REGION Network 5
   RUNG wire#powerrail
      { S7_Templates := "SrcType := Int" } EQ_Contact(in1 := #"BUFFER STATE", in2 := 0)
      I_Contact( #processing )
      I_Contact( #"MACHINE EXIT SENSOR" )
      I_Contact( #BUFFER_ITEMS_COUNT.QU )
      Move(in := 10, out1 => #"BUFFER STATE")
   END_RUNG
   // the same network as SCL:
   IF (#"BUFFER STATE" = 0) AND NOT #processing AND NOT #"MACHINE EXIT SENSOR" AND NOT #BUFFER_ITEMS_COUNT.QU THEN
       #"BUFFER STATE" := 10;
   END_IF;
END_REGION

REGION Network 6
   RUNG wire#powerrail
      #"ZONE 3 STOP BLADES LOGIC_Instance"("BUFFER STATE" := #"BUFFER STATE", "UP ELEVATOR STOP BLADE" => #"UP ELEVATOR STOP BLADE", "DOWN ELEVATOR STOP BLADE" => #"DOWN ELEVATOR STOP BLADE", "BRIDGE STOP BLADE 1" => #"BRIDGE STOP BLADE 1", "BRIDGE STOP BLADE 2" => #"BRIDGE STOP BLADE 2")
   END_RUNG
   // the same network as SCL:
   #"ZONE 3 STOP BLADES LOGIC_Instance"("BUFFER STATE" := #"BUFFER STATE",   // "ZONE 3 STOP BLADES LOGIC"
                           "UP ELEVATOR STOP BLADE" => #"UP ELEVATOR STOP BLADE",
                           "DOWN ELEVATOR STOP BLADE" => #"DOWN ELEVATOR STOP BLADE",
                           "BRIDGE STOP BLADE 1" => #"BRIDGE STOP BLADE 1",
                           "BRIDGE STOP BLADE 2" => #"BRIDGE STOP BLADE 2");
END_REGION

REGION Network 7
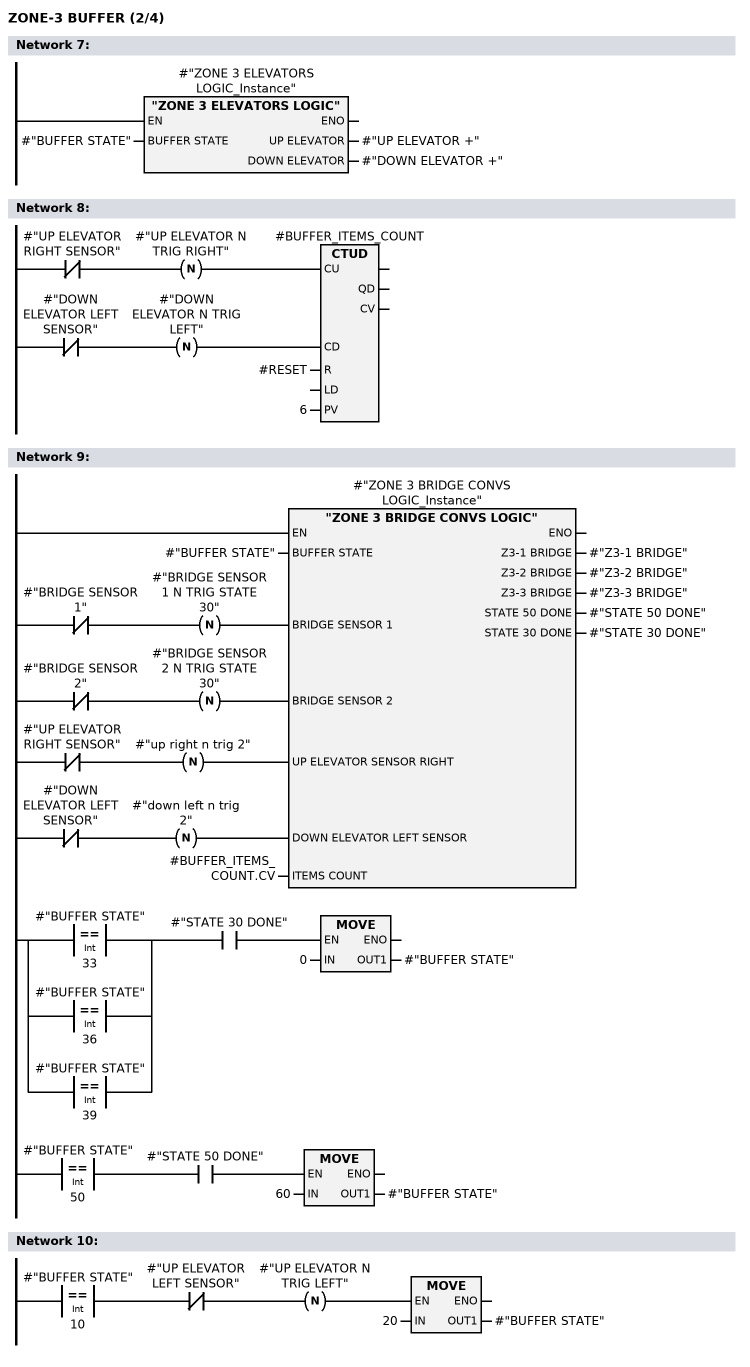
   RUNG wire#powerrail
      #"ZONE 3 ELEVATORS LOGIC_Instance"("BUFFER STATE" := #"BUFFER STATE", "UP ELEVATOR" => #"UP ELEVATOR +", "DOWN ELEVATOR" => #"DOWN ELEVATOR +")
   END_RUNG
   // the same network as SCL:
   #"ZONE 3 ELEVATORS LOGIC_Instance"("BUFFER STATE" := #"BUFFER STATE",   // "ZONE 3 ELEVATORS LOGIC"
                           "UP ELEVATOR" => #"UP ELEVATOR +",
                           "DOWN ELEVATOR" => #"DOWN ELEVATOR +");
END_REGION

REGION Network 8
   #_w1 := NOT (NOT #"UP ELEVATOR RIGHT SENSOR") AND #"UP ELEVATOR N TRIG RIGHT";   // falling edge
   #"UP ELEVATOR N TRIG RIGHT" := NOT #"UP ELEVATOR RIGHT SENSOR";
   #_w2 := NOT (NOT #"DOWN ELEVATOR LEFT SENSOR") AND #"DOWN ELEVATOR N TRIG LEFT";   // falling edge
   #"DOWN ELEVATOR N TRIG LEFT" := NOT #"DOWN ELEVATOR LEFT SENSOR";
   #BUFFER_ITEMS_COUNT(CU := #_w1, CD := #_w2, R := #RESET, PV := 6);   // CTUD
END_REGION

REGION Network 9
   RUNG wire#powerrail
      #"ZONE 3 BRIDGE CONVS LOGIC_Instance"("BRIDGE SENSOR 1" := wire#w1, "BRIDGE SENSOR 2" := wire#w2, "UP ELEVATOR SENSOR RIGHT" := wire#w3, "DOWN ELEVATOR LEFT SENSOR" := wire#w4, "BUFFER STATE" := #"BUFFER STATE", "ITEMS COUNT" := #BUFFER_ITEMS_COUNT.CV, "Z3-1 BRIDGE" => #"Z3-1 BRIDGE", "Z3-2 BRIDGE" => #"Z3-2 BRIDGE", "Z3-3 BRIDGE" => #"Z3-3 BRIDGE", "STATE 50 DONE" => #"STATE 50 DONE", "STATE 30 DONE" => #"STATE 30 DONE")
   END_RUNG
   RUNG wire#powerrail
      I_Contact( #"BRIDGE SENSOR 1" )
      N_Trig( #"BRIDGE SENSOR 1 N TRIG STATE 30" )
   END_RUNG wire#w1
   RUNG wire#powerrail
      I_Contact( #"BRIDGE SENSOR 2" )
      N_Trig( #"BRIDGE SENSOR 2 N TRIG STATE 30" )
   END_RUNG wire#w2
   RUNG wire#powerrail
      I_Contact( #"UP ELEVATOR RIGHT SENSOR" )
      N_Trig( #"up right n trig 2" )
   END_RUNG wire#w3
   RUNG wire#powerrail
      I_Contact( #"DOWN ELEVATOR LEFT SENSOR" )
      N_Trig( #"down left n trig 2" )
   END_RUNG wire#w4
   RUNG wire#powerrail
      { S7_Templates := "SrcType := Int" } EQ_Contact(in1 := #"BUFFER STATE", in2 := 33)
      wire#w5
      Contact( #"STATE 30 DONE" )
      Move(in := 0, out1 => #"BUFFER STATE")
   END_RUNG
   RUNG wire#powerrail
      { S7_Templates := "SrcType := Int" } EQ_Contact(in1 := #"BUFFER STATE", in2 := 36)
   END_RUNG wire#w5
   RUNG wire#powerrail
      { S7_Templates := "SrcType := Int" } EQ_Contact(in1 := #"BUFFER STATE", in2 := 39)
   END_RUNG wire#w5
   RUNG wire#powerrail
      { S7_Templates := "SrcType := Int" } EQ_Contact(in1 := #"BUFFER STATE", in2 := 50)
      Contact( #"STATE 50 DONE" )
      Move(in := 60, out1 => #"BUFFER STATE")
   END_RUNG
   // the same network as SCL:
   #_w1 := NOT (NOT #"BRIDGE SENSOR 1") AND #"BRIDGE SENSOR 1 N TRIG STATE 30";   // falling edge
   #"BRIDGE SENSOR 1 N TRIG STATE 30" := NOT #"BRIDGE SENSOR 1";
   #_w2 := NOT (NOT #"BRIDGE SENSOR 2") AND #"BRIDGE SENSOR 2 N TRIG STATE 30";   // falling edge
   #"BRIDGE SENSOR 2 N TRIG STATE 30" := NOT #"BRIDGE SENSOR 2";
   #_w3 := NOT (NOT #"UP ELEVATOR RIGHT SENSOR") AND #"up right n trig 2";   // falling edge
   #"up right n trig 2" := NOT #"UP ELEVATOR RIGHT SENSOR";
   #_w4 := NOT (NOT #"DOWN ELEVATOR LEFT SENSOR") AND #"down left n trig 2";   // falling edge
   #"down left n trig 2" := NOT #"DOWN ELEVATOR LEFT SENSOR";
   #"ZONE 3 BRIDGE CONVS LOGIC_Instance"("BUFFER STATE" := #"BUFFER STATE",   // "ZONE 3 BRIDGE CONVS LOGIC"
                           "BRIDGE SENSOR 1" := #_w1,
                           "BRIDGE SENSOR 2" := #_w2,
                           "UP ELEVATOR SENSOR RIGHT" := #_w3,
                           "DOWN ELEVATOR LEFT SENSOR" := #_w4,
                           "ITEMS COUNT" := #BUFFER_ITEMS_COUNT.CV,
                           "Z3-1 BRIDGE" => #"Z3-1 BRIDGE",
                           "Z3-2 BRIDGE" => #"Z3-2 BRIDGE",
                           "Z3-3 BRIDGE" => #"Z3-3 BRIDGE",
                           "STATE 50 DONE" => #"STATE 50 DONE",
                           "STATE 30 DONE" => #"STATE 30 DONE");
   IF ((#"BUFFER STATE" = 33) OR (#"BUFFER STATE" = 36) OR (#"BUFFER STATE" = 39)) AND #"STATE 30 DONE" THEN
       #"BUFFER STATE" := 0;
   END_IF;
   IF (#"BUFFER STATE" = 50) AND #"STATE 50 DONE" THEN #"BUFFER STATE" := 60; END_IF;
END_REGION

REGION Network 10
   RUNG wire#powerrail
      { S7_Templates := "SrcType := Int" } EQ_Contact(in1 := #"BUFFER STATE", in2 := 10)
      I_Contact( #"UP ELEVATOR LEFT SENSOR" )
      N_Trig( #"UP ELEVATOR N TRIG LEFT" )
      Move(in := 20, out1 => #"BUFFER STATE")
   END_RUNG
   // the same network as SCL:
   #_w1 := (#"BUFFER STATE" = 10) AND NOT #"UP ELEVATOR LEFT SENSOR";
   #_w2 := NOT #_w1 AND #"UP ELEVATOR N TRIG LEFT";   // falling edge
   #"UP ELEVATOR N TRIG LEFT" := #_w1;
   IF #_w2 THEN #"BUFFER STATE" := 20; END_IF;
END_REGION

REGION Network 11
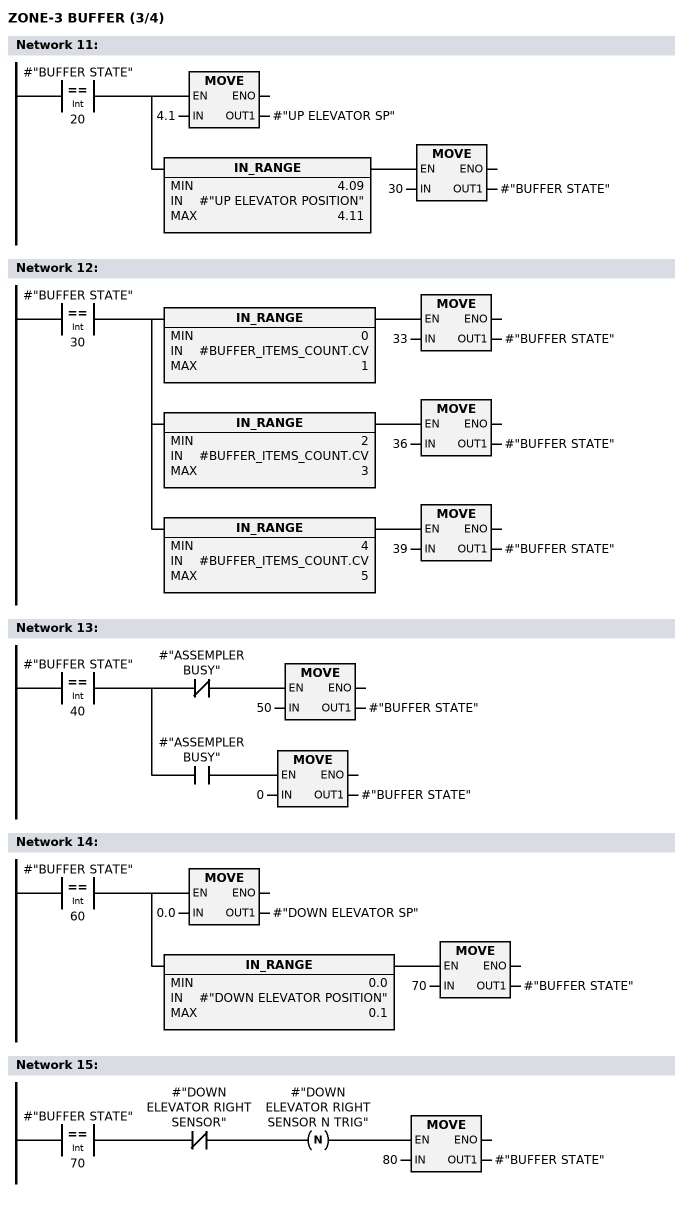
   RUNG wire#powerrail
      { S7_Templates := "SrcType := Int" } EQ_Contact(in1 := #"BUFFER STATE", in2 := 20)
      wire#w1
      Move(in := 4.1, out1 => #"UP ELEVATOR SP")
   END_RUNG
   RUNG wire#w1
      { S7_Templates := "SrcType := Real" } InRange(min := 4.09, in := #"UP ELEVATOR POSITION", max := 4.11)
      Move(in := 30, out1 => #"BUFFER STATE")
   END_RUNG
   // the same network as SCL:
   #_w1 := #"BUFFER STATE" = 20;
   IF #_w1 THEN #"UP ELEVATOR SP" := 4.1; END_IF;
   IF #_w1 AND (4.09 <= #"UP ELEVATOR POSITION") AND (#"UP ELEVATOR POSITION" <= 4.11) THEN
       #"BUFFER STATE" := 30;
   END_IF;
END_REGION

REGION Network 12
   RUNG wire#powerrail
      { S7_Templates := "SrcType := Int" } EQ_Contact(in1 := #"BUFFER STATE", in2 := 30)
      wire#w1
      { S7_Templates := "SrcType := Int" } InRange(min := 0, in := #BUFFER_ITEMS_COUNT.CV, max := 1)
      Move(in := 33, out1 => #"BUFFER STATE")
   END_RUNG
   RUNG wire#w1
      { S7_Templates := "SrcType := Int" } InRange(min := 2, in := #BUFFER_ITEMS_COUNT.CV, max := 3)
      Move(in := 36, out1 => #"BUFFER STATE")
   END_RUNG
   RUNG wire#w1
      { S7_Templates := "SrcType := Int" } InRange(min := 4, in := #BUFFER_ITEMS_COUNT.CV, max := 5)
      Move(in := 39, out1 => #"BUFFER STATE")
   END_RUNG
   // the same network as SCL:
   #_w1 := #"BUFFER STATE" = 30;
   IF #_w1 AND (0 <= #BUFFER_ITEMS_COUNT.CV) AND (#BUFFER_ITEMS_COUNT.CV <= 1) THEN
       #"BUFFER STATE" := 33;
   END_IF;
   IF #_w1 AND (2 <= #BUFFER_ITEMS_COUNT.CV) AND (#BUFFER_ITEMS_COUNT.CV <= 3) THEN
       #"BUFFER STATE" := 36;
   END_IF;
   IF #_w1 AND (4 <= #BUFFER_ITEMS_COUNT.CV) AND (#BUFFER_ITEMS_COUNT.CV <= 5) THEN
       #"BUFFER STATE" := 39;
   END_IF;
END_REGION

REGION Network 13
   RUNG wire#powerrail
      { S7_Templates := "SrcType := Int" } EQ_Contact(in1 := #"BUFFER STATE", in2 := 40)
      wire#w1
      I_Contact( #"ASSEMPLER BUSY" )
      Move(in := 50, out1 => #"BUFFER STATE")
   END_RUNG
   RUNG wire#w1
      Contact( #"ASSEMPLER BUSY" )
      Move(in := 0, out1 => #"BUFFER STATE")
   END_RUNG
   // the same network as SCL:
   #_w1 := #"BUFFER STATE" = 40;
   IF #_w1 AND NOT #"ASSEMPLER BUSY" THEN #"BUFFER STATE" := 50; END_IF;
   IF #_w1 AND #"ASSEMPLER BUSY" THEN #"BUFFER STATE" := 0; END_IF;
END_REGION

REGION Network 14
   RUNG wire#powerrail
      { S7_Templates := "SrcType := Int" } EQ_Contact(in1 := #"BUFFER STATE", in2 := 60)
      wire#w1
      Move(in := 0.0, out1 => #"DOWN ELEVATOR SP")
   END_RUNG
   RUNG wire#w1
      { S7_Templates := "SrcType := Real" } InRange(min := 0.0, in := #"DOWN ELEVATOR POSITION", max := 0.1)
      Move(in := 70, out1 => #"BUFFER STATE")
   END_RUNG
   // the same network as SCL:
   #_w1 := #"BUFFER STATE" = 60;
   IF #_w1 THEN #"DOWN ELEVATOR SP" := 0.0; END_IF;
   IF #_w1 AND (0.0 <= #"DOWN ELEVATOR POSITION") AND (#"DOWN ELEVATOR POSITION" <= 0.1) THEN
       #"BUFFER STATE" := 70;
   END_IF;
END_REGION

REGION Network 15
   RUNG wire#powerrail
      { S7_Templates := "SrcType := Int" } EQ_Contact(in1 := #"BUFFER STATE", in2 := 70)
      I_Contact( #"DOWN ELEVATOR RIGHT SENSOR" )
      N_Trig( #"DOWN ELEVATOR RIGHT SENSOR N TRIG" )
      Move(in := 80, out1 => #"BUFFER STATE")
   END_RUNG
   // the same network as SCL:
   #_w1 := (#"BUFFER STATE" = 70) AND NOT #"DOWN ELEVATOR RIGHT SENSOR";
   #_w2 := NOT #_w1 AND #"DOWN ELEVATOR RIGHT SENSOR N TRIG";   // falling edge
   #"DOWN ELEVATOR RIGHT SENSOR N TRIG" := #_w1;
   IF #_w2 THEN #"BUFFER STATE" := 80; END_IF;
END_REGION

REGION Network 16
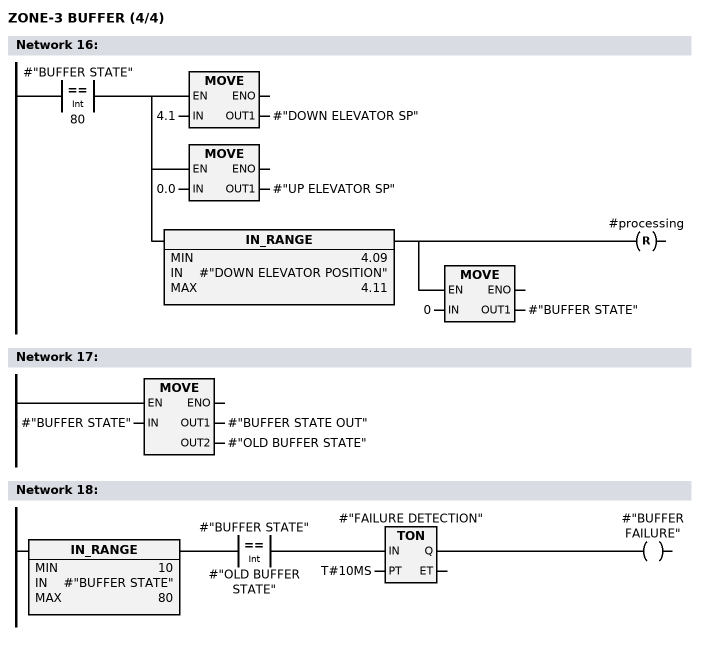
   RUNG wire#powerrail
      { S7_Templates := "SrcType := Int" } EQ_Contact(in1 := #"BUFFER STATE", in2 := 80)
      wire#w1
      Move(in := 4.1, out1 => #"DOWN ELEVATOR SP")
   END_RUNG
   RUNG wire#w1
      Move(in := 0.0, out1 => #"UP ELEVATOR SP")
   END_RUNG
   RUNG wire#w1
      { S7_Templates := "SrcType := Real" } InRange(min := 4.09, in := #"DOWN ELEVATOR POSITION", max := 4.11)
      wire#w2
      R_Coil( #processing )
   END_RUNG
   RUNG wire#w2
      Move(in := 0, out1 => #"BUFFER STATE")
   END_RUNG
   // the same network as SCL:
   #_w1 := #"BUFFER STATE" = 80;
   IF #_w1 THEN
       #"DOWN ELEVATOR SP" := 4.1;
       #"UP ELEVATOR SP" := 0.0;
   END_IF;
   IF #_w1 AND (4.09 <= #"DOWN ELEVATOR POSITION") AND (#"DOWN ELEVATOR POSITION" <= 4.11) THEN
       #processing := FALSE;
       #"BUFFER STATE" := 0;
   END_IF;
END_REGION

REGION Network 17
   RUNG wire#powerrail
      Move(in := #"BUFFER STATE", out1 => #"BUFFER STATE OUT", out2 => #"OLD BUFFER STATE")
   END_RUNG
   // the same network as SCL:
   #"BUFFER STATE OUT" := #"BUFFER STATE";
   #"OLD BUFFER STATE" := #"BUFFER STATE";
END_REGION

REGION Network 18
   #"FAILURE DETECTION"(IN := (10 <= #"BUFFER STATE") AND (#"BUFFER STATE" <= 80) AND (#"BUFFER STATE" = #"OLD BUFFER STATE"),   // TON
                        PT := T#10MS);
   #"BUFFER FAILURE" := #"FAILURE DETECTION".Q;
END_REGION
END_FUNCTION_BLOCK

FUNCTION_BLOCK "ZONE 3 ASSEMPLER"   // FB13, LAD
{ S7_Optimized_Access := 'TRUE' }
VERSION : 0.1
   VAR_INPUT
      EMERGENCY : Bool;
      "PRODUCT A AT ASSEMPLY" : Bool;
      "PRODUCT B AT ASSEMPLY" : Bool;
      "PRODUCT LEFT ASSEMPLY" : Bool;
      "POSITIONER A CLAMPED" : Bool;
      "POSITIONER B CLAMPED" : Bool;
      "POSITIONER B LIMIT" : Bool;
      "ASSEMPLER X POSITION" : Real;
      "ASSEMPLER Z POSITION'" : Real;
      "ITEM DETECTED" : Bool;
      "ASSEMPLER ROTATING" : Bool;
      "BUFFER A READY" : Bool;
      "BUFFER B READY" : Bool;
      RESET : Bool;
   END_VAR
   VAR_OUTPUT
      "POSITIONER A CLAMP" : Bool;
      "POSITIONER B CLAMP" : Bool;
      "POSITIONER B RAISE" : Bool;
      GRAP : Bool;
      ROTATE : Bool;
      "ROTATE CCW" : Bool;
      "X SET POINT" : Real;
      "Z SET POINT" : Real;
      "ASSEMPLER BUSY" : Bool;
      "ASSEMPER STATE OUT" : Int;
      "ASSEMPLER FAILURE" : Bool;
   END_VAR
   VAR
      "ASSEMPLER STATE" : Int;
      "POSITIONER LOGIC_Instance" : "POSITIONER LOGIC";
      "PRODUCT A N-TRIG" : Bool;
      "PRODUCT B N-TRIG" : Bool;
      "ASSEMPLER START" : Bool;
      "PRODUCT LEFT N TRIG" : Bool;
      "assempler rotation_Instance" : "assempler rotation";
      "TON-STATE-80-FAILURE" : TON_TIME;
      "MAINTENANCE MODE" : Bool;
      "MAINTENANCE P TRIG" : Bool;
      "MAINTENANCE N TRIG" : Bool;
      "ASSEMPLER SP MANAGMENT_Instance" : "ASSEMPLER SP MANAGMENT";
      "OLD STATE" : Int;
      "FAILURE DETECTION" : TON_TIME;
   END_VAR
   VAR_TEMP   // added for the SCL form of the ladder/FBD networks
      _w1 : Bool;
      _w2 : Bool;
   END_VAR
BEGIN

REGION Network 1
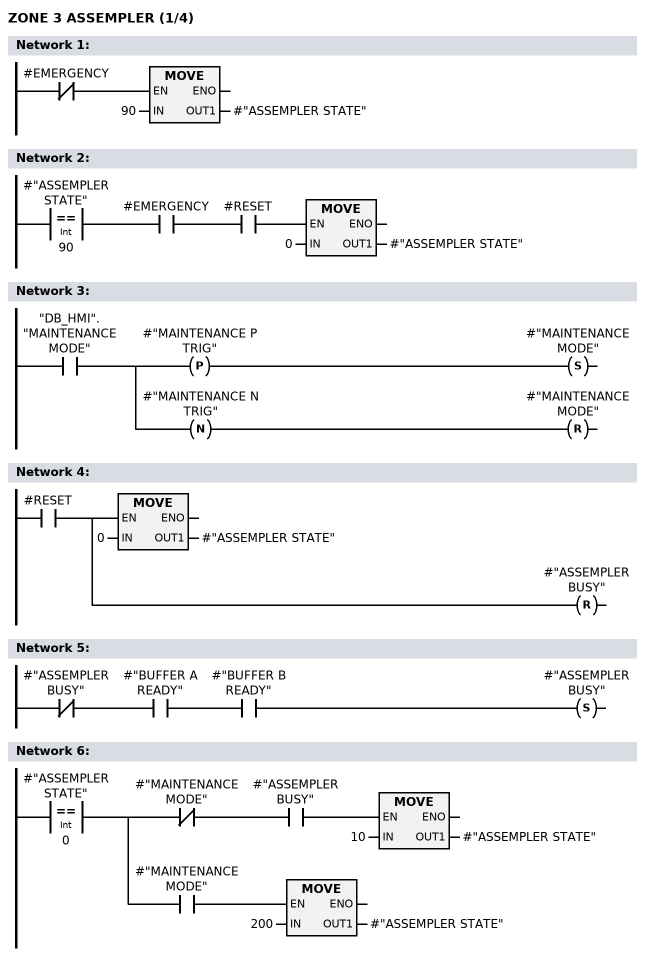
   RUNG wire#powerrail
      I_Contact( #EMERGENCY )
      Move(in := 90, out1 => #"ASSEMPLER STATE")
   END_RUNG
   // the same network as SCL:
   IF NOT #EMERGENCY THEN #"ASSEMPLER STATE" := 90; END_IF;
END_REGION

REGION Network 2
   RUNG wire#powerrail
      { S7_Templates := "SrcType := Int" } EQ_Contact(in1 := #"ASSEMPLER STATE", in2 := 90)
      Contact( #EMERGENCY )
      Contact( #RESET )
      Move(in := 0, out1 => #"ASSEMPLER STATE")
   END_RUNG
   // the same network as SCL:
   IF (#"ASSEMPLER STATE" = 90) AND #EMERGENCY AND #RESET THEN #"ASSEMPLER STATE" := 0; END_IF;
END_REGION

REGION Network 3
   RUNG wire#powerrail
      Contact( "DB_HMI"."MAINTENANCE MODE" )
      wire#w1
      P_Trig( #"MAINTENANCE P TRIG" )
      S_Coil( #"MAINTENANCE MODE" )
   END_RUNG
   RUNG wire#w1
      N_Trig( #"MAINTENANCE N TRIG" )
      R_Coil( #"MAINTENANCE MODE" )
   END_RUNG
   // the same network as SCL:
   #_w1 := "DB_HMI"."MAINTENANCE MODE" AND NOT #"MAINTENANCE P TRIG";   // rising edge
   #"MAINTENANCE P TRIG" := "DB_HMI"."MAINTENANCE MODE";
   IF #_w1 THEN #"MAINTENANCE MODE" := TRUE; END_IF;
   #_w2 := NOT "DB_HMI"."MAINTENANCE MODE" AND #"MAINTENANCE N TRIG";   // falling edge
   #"MAINTENANCE N TRIG" := "DB_HMI"."MAINTENANCE MODE";
   IF #_w2 THEN #"MAINTENANCE MODE" := FALSE; END_IF;
END_REGION

REGION Network 4
   RUNG wire#powerrail
      Contact( #RESET )
      wire#w1
      Move(in := 0, out1 => #"ASSEMPLER STATE")
   END_RUNG
   RUNG wire#w1
      R_Coil( #"ASSEMPLER BUSY" )
   END_RUNG
   // the same network as SCL:
   IF #RESET THEN
       #"ASSEMPLER STATE" := 0;
       #"ASSEMPLER BUSY" := FALSE;
   END_IF;
END_REGION

REGION Network 5
   RUNG wire#powerrail
      I_Contact( #"ASSEMPLER BUSY" )
      Contact( #"BUFFER A READY" )
      Contact( #"BUFFER B READY" )
      S_Coil( #"ASSEMPLER BUSY" )
   END_RUNG
   // the same network as SCL:
   IF NOT #"ASSEMPLER BUSY" AND #"BUFFER A READY" AND #"BUFFER B READY" THEN
       #"ASSEMPLER BUSY" := TRUE;
   END_IF;
END_REGION

REGION Network 6
   RUNG wire#powerrail
      { S7_Templates := "SrcType := Int" } EQ_Contact(in1 := #"ASSEMPLER STATE", in2 := 0)
      wire#w1
      I_Contact( #"MAINTENANCE MODE" )
      Contact( #"ASSEMPLER BUSY" )
      Move(in := 10, out1 => #"ASSEMPLER STATE")
   END_RUNG
   RUNG wire#w1
      Contact( #"MAINTENANCE MODE" )
      Move(in := 200, out1 => #"ASSEMPLER STATE")
   END_RUNG
   // the same network as SCL:
   #_w1 := #"ASSEMPLER STATE" = 0;
   IF #_w1 AND NOT #"MAINTENANCE MODE" AND #"ASSEMPLER BUSY" THEN #"ASSEMPLER STATE" := 10; END_IF;
   IF #_w1 AND #"MAINTENANCE MODE" THEN #"ASSEMPLER STATE" := 200; END_IF;
END_REGION

REGION Network 7
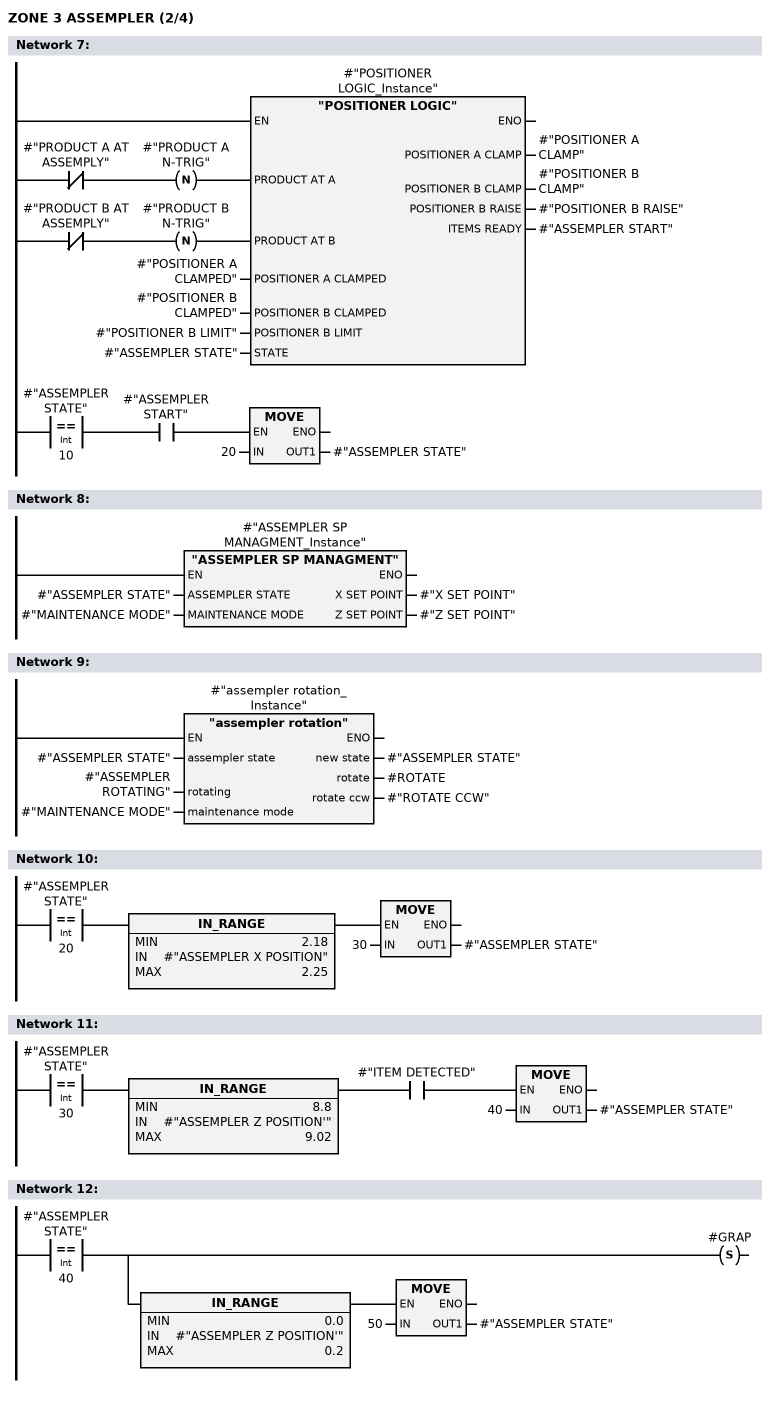
   RUNG wire#powerrail
      #"POSITIONER LOGIC_Instance"("PRODUCT AT A" := wire#w1, "PRODUCT AT B" := wire#w2, "POSITIONER A CLAMPED" := #"POSITIONER A CLAMPED", "POSITIONER B CLAMPED" := #"POSITIONER B CLAMPED", "POSITIONER B LIMIT" := #"POSITIONER B LIMIT", STATE := #"ASSEMPLER STATE", "POSITIONER A CLAMP" => #"POSITIONER A CLAMP", "POSITIONER B CLAMP" => #"POSITIONER B CLAMP", "POSITIONER B RAISE" => #"POSITIONER B RAISE", "ITEMS READY" => #"ASSEMPLER START")
   END_RUNG
   RUNG wire#powerrail
      I_Contact( #"PRODUCT A AT ASSEMPLY" )
      N_Trig( #"PRODUCT A N-TRIG" )
   END_RUNG wire#w1
   RUNG wire#powerrail
      I_Contact( #"PRODUCT B AT ASSEMPLY" )
      N_Trig( #"PRODUCT B N-TRIG" )
   END_RUNG wire#w2
   RUNG wire#powerrail
      { S7_Templates := "SrcType := Int" } EQ_Contact(in1 := #"ASSEMPLER STATE", in2 := 10)
      Contact( #"ASSEMPLER START" )
      Move(in := 20, out1 => #"ASSEMPLER STATE")
   END_RUNG
   // the same network as SCL:
   #_w1 := NOT (NOT #"PRODUCT A AT ASSEMPLY") AND #"PRODUCT A N-TRIG";   // falling edge
   #"PRODUCT A N-TRIG" := NOT #"PRODUCT A AT ASSEMPLY";
   #_w2 := NOT (NOT #"PRODUCT B AT ASSEMPLY") AND #"PRODUCT B N-TRIG";   // falling edge
   #"PRODUCT B N-TRIG" := NOT #"PRODUCT B AT ASSEMPLY";
   #"POSITIONER LOGIC_Instance"("PRODUCT AT A" := #_w1,   // "POSITIONER LOGIC"
                           "PRODUCT AT B" := #_w2,
                           "POSITIONER A CLAMPED" := #"POSITIONER A CLAMPED",
                           "POSITIONER B CLAMPED" := #"POSITIONER B CLAMPED",
                           "POSITIONER B LIMIT" := #"POSITIONER B LIMIT",
                           STATE := #"ASSEMPLER STATE",
                           "POSITIONER A CLAMP" => #"POSITIONER A CLAMP",
                           "POSITIONER B CLAMP" => #"POSITIONER B CLAMP",
                           "POSITIONER B RAISE" => #"POSITIONER B RAISE",
                           "ITEMS READY" => #"ASSEMPLER START");
   IF (#"ASSEMPLER STATE" = 10) AND #"ASSEMPLER START" THEN #"ASSEMPLER STATE" := 20; END_IF;
END_REGION

REGION Network 8
   RUNG wire#powerrail
      #"ASSEMPLER SP MANAGMENT_Instance"("ASSEMPLER STATE" := #"ASSEMPLER STATE", "MAINTENANCE MODE" := #"MAINTENANCE MODE", "X SET POINT" => #"X SET POINT", "Z SET POINT" => #"Z SET POINT")
   END_RUNG
   // the same network as SCL:
   #"ASSEMPLER SP MANAGMENT_Instance"("ASSEMPLER STATE" := #"ASSEMPLER STATE",   // "ASSEMPLER SP MANAGMENT"
                           "MAINTENANCE MODE" := #"MAINTENANCE MODE",
                           "X SET POINT" => #"X SET POINT",
                           "Z SET POINT" => #"Z SET POINT");
END_REGION

REGION Network 9
   RUNG wire#powerrail
      #"assempler rotation_Instance"("assempler state" := #"ASSEMPLER STATE", rotating := #"ASSEMPLER ROTATING", "maintenance mode" := #"MAINTENANCE MODE", "new state" => #"ASSEMPLER STATE", rotate => #ROTATE, "rotate ccw" => #"ROTATE CCW")
   END_RUNG
   // the same network as SCL:
   #"assempler rotation_Instance"("assempler state" := #"ASSEMPLER STATE",   // "assempler rotation"
                           rotating := #"ASSEMPLER ROTATING",
                           "maintenance mode" := #"MAINTENANCE MODE",
                           "new state" => #"ASSEMPLER STATE",
                           rotate => #ROTATE,
                           "rotate ccw" => #"ROTATE CCW");
END_REGION

REGION Network 10
   RUNG wire#powerrail
      { S7_Templates := "SrcType := Int" } EQ_Contact(in1 := #"ASSEMPLER STATE", in2 := 20)
      { S7_Templates := "SrcType := Real" } InRange(min := 2.18, in := #"ASSEMPLER X POSITION", max := 2.25)
      Move(in := 30, out1 => #"ASSEMPLER STATE")
   END_RUNG
   // the same network as SCL:
   IF (#"ASSEMPLER STATE" = 20) AND (2.18 <= #"ASSEMPLER X POSITION") AND (#"ASSEMPLER X POSITION" <= 2.25) THEN
       #"ASSEMPLER STATE" := 30;
   END_IF;
END_REGION

REGION Network 11
   RUNG wire#powerrail
      { S7_Templates := "SrcType := Int" } EQ_Contact(in1 := #"ASSEMPLER STATE", in2 := 30)
      { S7_Templates := "SrcType := Real" } InRange(min := 8.8, in := #"ASSEMPLER Z POSITION'", max := 9.02)
      Contact( #"ITEM DETECTED" )
      Move(in := 40, out1 => #"ASSEMPLER STATE")
   END_RUNG
   // the same network as SCL:
   IF (#"ASSEMPLER STATE" = 30) AND (8.8 <= #"ASSEMPLER Z POSITION'") AND (#"ASSEMPLER Z POSITION'" <= 9.02) AND #"ITEM DETECTED" THEN
       #"ASSEMPLER STATE" := 40;
   END_IF;
END_REGION

REGION Network 12
   RUNG wire#powerrail
      { S7_Templates := "SrcType := Int" } EQ_Contact(in1 := #"ASSEMPLER STATE", in2 := 40)
      wire#w1
      S_Coil( #GRAP )
   END_RUNG
   RUNG wire#w1
      { S7_Templates := "SrcType := Real" } InRange(min := 0.0, in := #"ASSEMPLER Z POSITION'", max := 0.2)
      Move(in := 50, out1 => #"ASSEMPLER STATE")
   END_RUNG
   // the same network as SCL:
   #_w1 := #"ASSEMPLER STATE" = 40;
   IF #_w1 THEN #GRAP := TRUE; END_IF;
   IF #_w1 AND (0.0 <= #"ASSEMPLER Z POSITION'") AND (#"ASSEMPLER Z POSITION'" <= 0.2) THEN
       #"ASSEMPLER STATE" := 50;
   END_IF;
END_REGION

REGION Network 13
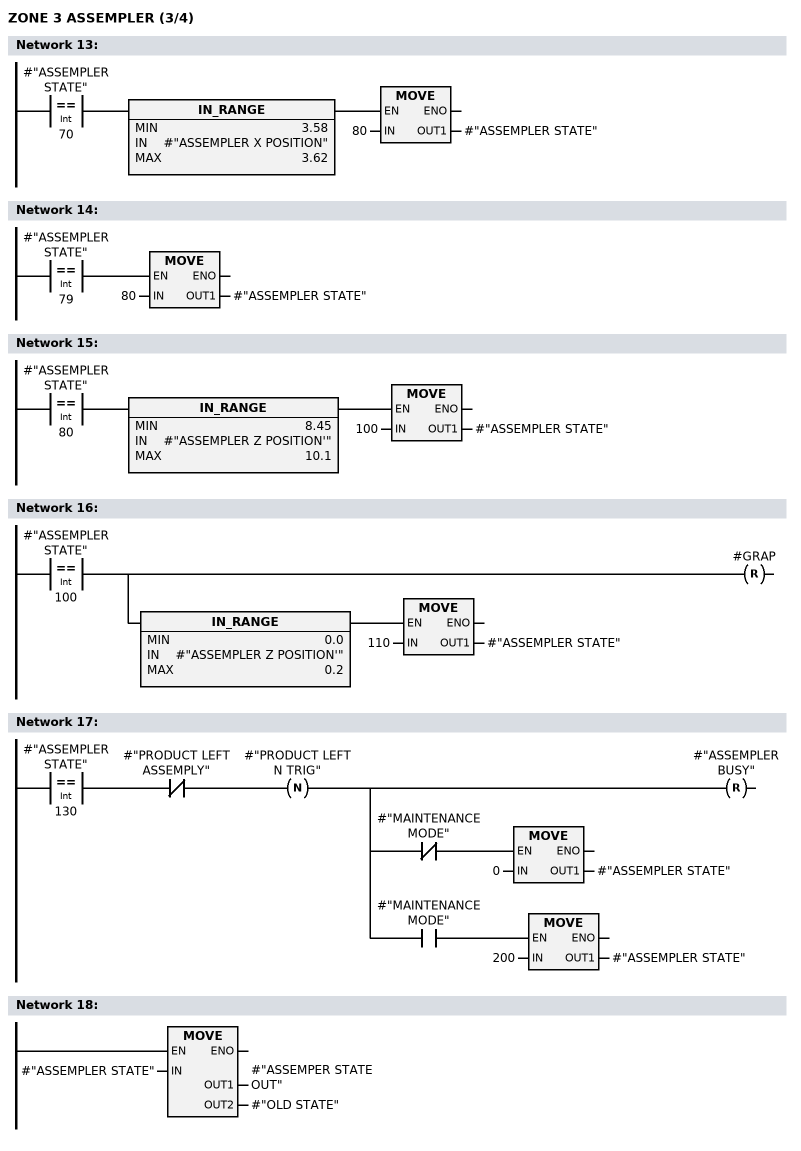
   RUNG wire#powerrail
      { S7_Templates := "SrcType := Int" } EQ_Contact(in1 := #"ASSEMPLER STATE", in2 := 70)
      { S7_Templates := "SrcType := Real" } InRange(min := 3.58, in := #"ASSEMPLER X POSITION", max := 3.62)
      Move(in := 80, out1 => #"ASSEMPLER STATE")
   END_RUNG
   // the same network as SCL:
   IF (#"ASSEMPLER STATE" = 70) AND (3.58 <= #"ASSEMPLER X POSITION") AND (#"ASSEMPLER X POSITION" <= 3.62) THEN
       #"ASSEMPLER STATE" := 80;
   END_IF;
END_REGION

REGION Network 14
   RUNG wire#powerrail
      { S7_Templates := "SrcType := Int" } EQ_Contact(in1 := #"ASSEMPLER STATE", in2 := 79)
      Move(in := 80, out1 => #"ASSEMPLER STATE")
   END_RUNG
   // the same network as SCL:
   IF #"ASSEMPLER STATE" = 79 THEN #"ASSEMPLER STATE" := 80; END_IF;
END_REGION

REGION Network 15
   RUNG wire#powerrail
      { S7_Templates := "SrcType := Int" } EQ_Contact(in1 := #"ASSEMPLER STATE", in2 := 80)
      { S7_Templates := "SrcType := Real" } InRange(min := 8.45, in := #"ASSEMPLER Z POSITION'", max := 10.1)
      Move(in := 100, out1 => #"ASSEMPLER STATE")
   END_RUNG
   // the same network as SCL:
   IF (#"ASSEMPLER STATE" = 80) AND (8.45 <= #"ASSEMPLER Z POSITION'") AND (#"ASSEMPLER Z POSITION'" <= 10.1) THEN
       #"ASSEMPLER STATE" := 100;
   END_IF;
END_REGION

REGION Network 16
   RUNG wire#powerrail
      { S7_Templates := "SrcType := Int" } EQ_Contact(in1 := #"ASSEMPLER STATE", in2 := 100)
      wire#w1
      R_Coil( #GRAP )
   END_RUNG
   RUNG wire#w1
      { S7_Templates := "SrcType := Real" } InRange(min := 0.0, in := #"ASSEMPLER Z POSITION'", max := 0.2)
      Move(in := 110, out1 => #"ASSEMPLER STATE")
   END_RUNG
   // the same network as SCL:
   #_w1 := #"ASSEMPLER STATE" = 100;
   IF #_w1 THEN #GRAP := FALSE; END_IF;
   IF #_w1 AND (0.0 <= #"ASSEMPLER Z POSITION'") AND (#"ASSEMPLER Z POSITION'" <= 0.2) THEN
       #"ASSEMPLER STATE" := 110;
   END_IF;
END_REGION

REGION Network 17
   RUNG wire#powerrail
      { S7_Templates := "SrcType := Int" } EQ_Contact(in1 := #"ASSEMPLER STATE", in2 := 130)
      I_Contact( #"PRODUCT LEFT ASSEMPLY" )
      N_Trig( #"PRODUCT LEFT N TRIG" )
      wire#w1
      R_Coil( #"ASSEMPLER BUSY" )
   END_RUNG
   RUNG wire#w1
      I_Contact( #"MAINTENANCE MODE" )
      Move(in := 0, out1 => #"ASSEMPLER STATE")
   END_RUNG
   RUNG wire#w1
      Contact( #"MAINTENANCE MODE" )
      Move(in := 200, out1 => #"ASSEMPLER STATE")
   END_RUNG
   // the same network as SCL:
   #_w1 := (#"ASSEMPLER STATE" = 130) AND NOT #"PRODUCT LEFT ASSEMPLY";
   #_w2 := NOT #_w1 AND #"PRODUCT LEFT N TRIG";   // falling edge
   #"PRODUCT LEFT N TRIG" := #_w1;
   IF #_w2 THEN #"ASSEMPLER BUSY" := FALSE; END_IF;
   IF #_w2 AND NOT #"MAINTENANCE MODE" THEN #"ASSEMPLER STATE" := 0; END_IF;
   IF #_w2 AND #"MAINTENANCE MODE" THEN #"ASSEMPLER STATE" := 200; END_IF;
END_REGION

REGION Network 18
   RUNG wire#powerrail
      Move(in := #"ASSEMPLER STATE", out1 => #"ASSEMPER STATE OUT", out2 => #"OLD STATE")
   END_RUNG
   // the same network as SCL:
   #"ASSEMPER STATE OUT" := #"ASSEMPLER STATE";
   #"OLD STATE" := #"ASSEMPLER STATE";
END_REGION

REGION Network 19
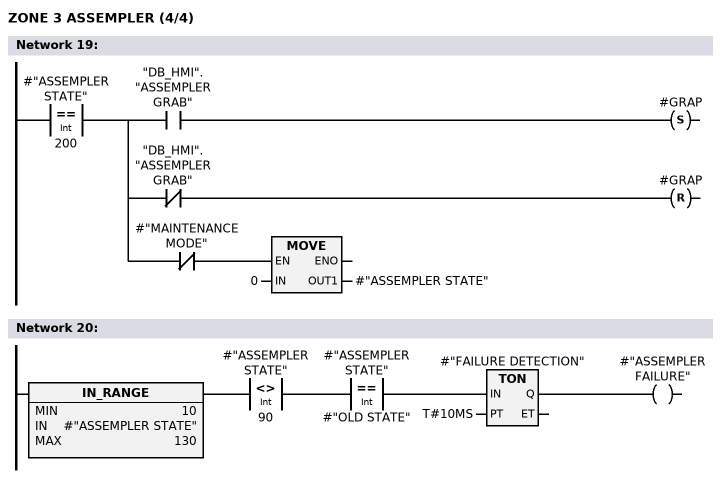
   RUNG wire#powerrail
      { S7_Templates := "SrcType := Int" } EQ_Contact(in1 := #"ASSEMPLER STATE", in2 := 200)
      wire#w1
      Contact( "DB_HMI"."ASSEMPLER GRAB" )
      S_Coil( #GRAP )
   END_RUNG
   RUNG wire#w1
      I_Contact( "DB_HMI"."ASSEMPLER GRAB" )
      R_Coil( #GRAP )
   END_RUNG
   RUNG wire#w1
      I_Contact( #"MAINTENANCE MODE" )
      Move(in := 0, out1 => #"ASSEMPLER STATE")
   END_RUNG
   // the same network as SCL:
   #_w1 := #"ASSEMPLER STATE" = 200;
   IF #_w1 AND "DB_HMI"."ASSEMPLER GRAB" THEN #GRAP := TRUE; END_IF;
   IF #_w1 AND NOT "DB_HMI"."ASSEMPLER GRAB" THEN #GRAP := FALSE; END_IF;
   IF #_w1 AND NOT #"MAINTENANCE MODE" THEN #"ASSEMPLER STATE" := 0; END_IF;
END_REGION

REGION Network 20
   #"FAILURE DETECTION"(IN := (10 <= #"ASSEMPLER STATE") AND (#"ASSEMPLER STATE" <= 130) AND (#"ASSEMPLER STATE" <> 90) AND (#"ASSEMPLER STATE" = #"OLD STATE"),   // TON
                        PT := T#10MS);
   #"ASSEMPLER FAILURE" := #"FAILURE DETECTION".Q;
END_REGION
END_FUNCTION_BLOCK

// folder: Zone_3_blocks/ASSEMPLER SUB BLOCKS

FUNCTION_BLOCK "assempler rotation"   // FB14, SCL
{ S7_Optimized_Access := 'TRUE' }
VERSION : 0.1
   VAR_INPUT
      "assempler state" : Int;
      rotating : Bool;
      "maintenance mode" : Bool;
   END_VAR
   VAR_OUTPUT
      "new state" : Int;
      rotate : Bool;
      "rotate ccw" : Bool;
   END_VAR
   VAR
      "TON-0" : TON_TIME;
      done : Bool;
      "TON-1" : TON_TIME;
      advance : Bool;
      cooldown : Bool;
      "ton-3" : TON_TIME;
      done2 : Bool;
      cooldown2 : Bool;
      advance2 : Bool;
      "ton-4" : TON_TIME;
   END_VAR
BEGIN
   #"TON-0"(IN := #rotate,
                PT := T#500ms,
                Q => #done);
   #"TON-1"(IN:=#cooldown,
            PT:=T#500ms,
            Q=>#advance);
   #"ton-3"(IN := #"rotate ccw",
            PT := T#500ms,
            Q => #done2);
   #"ton-4"(IN := #cooldown2,
            PT := T#500ms,
            Q => #advance2);


   IF #"maintenance mode" AND #"assempler state" = 200 THEN
       #"new state" := 200;
       IF "DB_HMI"."ASSEMPLER ROT CW" THEN
           #rotate := 1;
           IF #done THEN
               #rotate := 0;
               #cooldown := 1;
               IF #advance THEN
                   #cooldown := 0;
                   "DB_HMI"."ASSEMPLER ROT CW" := 0;
               END_IF;
           END_IF;
       END_IF;
       IF "DB_HMI"."ASSEMPLER ROT CCW" THEN
           #"rotate ccw" := 1;
           IF #done2 THEN
               #"rotate ccw":= 0;
               #cooldown2 := 1;
               IF #advance2 THEN
                   #cooldown := 0;
                   "DB_HMI"."ASSEMPLER ROT CCW" := 0;
               END_IF;
           END_IF;
       END_IF;
   ELSE

       CASE #"assempler state" OF
           50:
               #rotate := 1;
               IF #done THEN

                   #rotate := 0;
                   #cooldown := 1;
                   IF #advance THEN
                       #"new state" := 60;
                       #cooldown := 0;
                   END_IF;
               END_IF;
           60:
               #rotate := 1;
               IF #done THEN
                   #rotate := 0;
                   #cooldown := 1;
                   IF #advance THEN
                       #"new state" := 70;
                       #cooldown := 0;
                   END_IF;
               END_IF;
           110:
               #rotate := 1;
               IF #done THEN
                   #rotate := 0;
                   #cooldown := 1;
                   IF #advance THEN
                       #"new state" := 120;
                       #cooldown := 0;
                   END_IF;
               END_IF;
           120:
               #rotate := 1;
               IF #done THEN
                   #rotate := 0;
                   #cooldown := 1;
                   IF #advance THEN
                       #"new state" := 130;
                       #cooldown := 0;
                   END_IF;
               END_IF;

           ELSE
               #"new state" := #"assempler state";
       END_CASE;
   END_IF;
END_FUNCTION_BLOCK

FUNCTION_BLOCK "POSITIONER LOGIC"   // FB15, SCL
{ S7_Optimized_Access := 'TRUE' }
VERSION : 0.1
   VAR_INPUT
      "PRODUCT AT A" : Bool;
      "PRODUCT AT B" : Bool;
      "POSITIONER A CLAMPED" : Bool;
      "POSITIONER B CLAMPED" : Bool;
      "POSITIONER B LIMIT" : Bool;
      STATE : Int;
   END_VAR
   VAR_OUTPUT
      "POSITIONER A CLAMP" : Bool;
      "POSITIONER B CLAMP" : Bool;
      "POSITIONER B RAISE" : Bool;
      "ITEMS READY" : Bool;
   END_VAR
   VAR
      "AT  A" : Bool;
      "AT B" : Bool;
   END_VAR
BEGIN
   IF #"PRODUCT AT A" THEN
       #"AT  A" := 1;
   END_IF;
   IF #"PRODUCT AT B" THEN
       #"AT B" := 1;
   END_IF;
   CASE #STATE OF
       0:
           #"POSITIONER A CLAMP" := 0;
           #"POSITIONER B CLAMP" := 0;
           #"AT  A" := 0;
           #"AT B" := 0;
       10:
           #"POSITIONER B RAISE" := 0;
           IF #"AT  A" THEN
               #"POSITIONER A CLAMP" := 1;
           ELSE
               #"POSITIONER A CLAMP" := 0;
           END_IF;
           IF #"AT B" THEN
               #"POSITIONER B CLAMP" := 1;
           ELSE
               #"POSITIONER B CLAMP" := 0;
           END_IF;
           IF #"POSITIONER A CLAMPED" AND #"POSITIONER B CLAMPED" THEN
               #"ITEMS READY" := 1;
           END_IF;

       40:  
           #"POSITIONER A CLAMP" := 0;
           #"ITEMS READY" := 0;
           #"POSITIONER B RAISE" := 0;
       100:
           #"POSITIONER B CLAMP" := 0;
           #"ITEMS READY" := 0;
           #"POSITIONER B RAISE" := 0;
       130:
           #"POSITIONER B RAISE" := 1;
           #"ITEMS READY" := 0;
           #"AT  A" := 0;
           #"AT B" := 0;
       90:
           #"POSITIONER A CLAMP" := 0;
           #"POSITIONER B CLAMP" := 0;
           #"AT  A" := 0;
           #"AT B" := 0;
           #"ITEMS READY" := 0;
           #"POSITIONER B RAISE" := 0;
       ELSE  
           #"ITEMS READY" := 0;
           #"POSITIONER B RAISE" := 0;

   END_CASE;
END_FUNCTION_BLOCK

FUNCTION_BLOCK "ASSEMPLER SP MANAGMENT"   // FB23, SCL
{ S7_Optimized_Access := 'TRUE' }
VERSION : 0.1
   VAR_INPUT
      "ASSEMPLER STATE" : Int;
      "MAINTENANCE MODE" : Bool;
   END_VAR
   VAR_OUTPUT
      "X SET POINT" : Real;
      "Z SET POINT" : Real;
   END_VAR
BEGIN
   IF #"MAINTENANCE MODE" AND #"ASSEMPLER STATE"=200 THEN
       #"X SET POINT" := "DB_HMI"."ASSEMPLER X";
       #"Z SET POINT" := "DB_HMI"."ASSEMPLER Z";
   ELSE
       CASE #"ASSEMPLER STATE" OF
           0:
               #"X SET POINT" := 0.0;
               #"Z SET POINT" := 0.0;
           10:
               #"X SET POINT" := 0.0;
               #"Z SET POINT" := 0.0;
           20:
               #"X SET POINT" := 2.2;
               #"Z SET POINT" := 0.0;
           30:
               #"X SET POINT" := 2.2;
               #"Z SET POINT" := 9.0;
           40..60:
               #"X SET POINT" := 2.2;
               #"Z SET POINT" := 0.0;
           70:
               #"X SET POINT" := 3.6;
               #"Z SET POINT" := 0.0;
           79:
               #"X SET POINT" := 3.3;
           80:
               #"Z SET POINT" := 10.0;
           100:
               #"Z SET POINT" := 0.0;
           90:
               #"X SET POINT" := 0.0;
               #"Z SET POINT" := 0.0;


           ELSE  
               #"X SET POINT" := 0.0;
               #"Z SET POINT" := 0.0;
       END_CASE;
   END_IF;
END_FUNCTION_BLOCK

// folder: Zone_3_blocks/BUFFER SUB BLOCKS

FUNCTION_BLOCK "ZONE 3 STOP BLADES LOGIC"   // FB9, SCL
{ S7_Optimized_Access := 'TRUE' }
VERSION : 0.1
   VAR_INPUT
      "BUFFER STATE" : Int;
   END_VAR
   VAR_OUTPUT
      "UP ELEVATOR STOP BLADE" : Bool;
      "DOWN ELEVATOR STOP BLADE" : Bool;
      "BRIDGE STOP BLADE 1" : Bool;
      "BRIDGE STOP BLADE 2" : Bool;
   END_VAR
BEGIN
   CASE #"BUFFER STATE" OF
       10:  
           #"UP ELEVATOR STOP BLADE" := 0;
           #"DOWN ELEVATOR STOP BLADE" := 1;
           #"BRIDGE STOP BLADE 1" := 1;
           #"BRIDGE STOP BLADE 2" := 1;
       20:  
           #"UP ELEVATOR STOP BLADE" := 1;
           #"DOWN ELEVATOR STOP BLADE" := 1;
           #"BRIDGE STOP BLADE 1" := 1;
           #"BRIDGE STOP BLADE 2" := 1;
       30:
           #"UP ELEVATOR STOP BLADE" := 1;
           #"DOWN ELEVATOR STOP BLADE" := 1;
           #"BRIDGE STOP BLADE 1" := 1;
           #"BRIDGE STOP BLADE 2" := 1;

       33:
           #"UP ELEVATOR STOP BLADE" := 1;
           #"DOWN ELEVATOR STOP BLADE" := 1;
           #"BRIDGE STOP BLADE 1" := 0;
           #"BRIDGE STOP BLADE 2" := 0;
       36:
           #"UP ELEVATOR STOP BLADE" := 1;
           #"DOWN ELEVATOR STOP BLADE" := 1;
           #"BRIDGE STOP BLADE 1" := 0;
           #"BRIDGE STOP BLADE 2" := 1;
       39:
           #"UP ELEVATOR STOP BLADE" := 1;
           #"DOWN ELEVATOR STOP BLADE" := 1;
           #"BRIDGE STOP BLADE 1" := 1;
           #"BRIDGE STOP BLADE 2" := 1;
       40:
           #"UP ELEVATOR STOP BLADE" := 1;
           #"DOWN ELEVATOR STOP BLADE" := 0;
           #"BRIDGE STOP BLADE 1" := 1;
           #"BRIDGE STOP BLADE 2" := 1;
       50:
           #"UP ELEVATOR STOP BLADE" := 1;
           #"DOWN ELEVATOR STOP BLADE" := 0;
           #"BRIDGE STOP BLADE 1" := 0;
           #"BRIDGE STOP BLADE 2" := 0;
       60:
           #"UP ELEVATOR STOP BLADE" := 1;
           #"DOWN ELEVATOR STOP BLADE" := 1;
           #"BRIDGE STOP BLADE 1" := 1;
           #"BRIDGE STOP BLADE 2" := 1;
       ELSE  // Statement section ELSE
           #"UP ELEVATOR STOP BLADE" := 1;
           #"DOWN ELEVATOR STOP BLADE" := 1;
           #"BRIDGE STOP BLADE 1" := 1;
           #"BRIDGE STOP BLADE 2" := 1;
   END_CASE;
END_FUNCTION_BLOCK

FUNCTION_BLOCK "ZONE 3 ADVANCING THE BUFFER"   // FB10, SCL
{ S7_Optimized_Access := 'TRUE' }